   "14_DQ_Data_24PF2" : Bool = PLC "14_DQ_Data".24PF2 AT %DB1.DBX0.0, 1 s
   "19_AUTO_CMNDS_Data_PIT402_Target" : Real = PLC "19_AUTO_CMNDS_Data".PIT402_Target AT %DB1.DBD0, 1 s
   "80_From_HMI_RST_E500A_RT" : Bool = PLC "80_From_HMI".RST_E500A_RT AT %DB1.DBX0.0, 1 s
   "10_DI_Data_CV312_OPN" : Bool = PLC "10_DI_Data".CV312_OPN AT %DB1.DBX0.0, 1 s
   "10_DI_Data_CV312_CLSD" : Bool = PLC "10_DI_Data".CV312_CLSD AT %DB1.DBX0.0, 1 s
   "Clock_1Hz" : Bool = PLC Clock_1Hz AT %M0.5, 500 ms
   "14_DQ_Data_24K3(1)" : Bool = PLC "14_DQ_Data".24K3 AT %DB1.DBX0.0, 1 s
   "12_AI_Data_LIT305_SCALED" : Real = PLC "12_AI_Data".LIT305_SCALED AT %DB1.DBX0.0, 1 s
   "80_From_HMI_BWT_BYPASS(1)" : Bool = PLC "80_From_HMI".BWT_BYPASS AT %DB1.DBX0.0, 1 s
   "80_From_HMI_CRG_BLNK_MODE(1)" : Bool = PLC "80_From_HMI".CRG_BLNK_MODE AT %DB1.DBX0.0, 1 s
   "80_From_HMI_BWT_BYPASS" : Bool = PLC "80_From_HMI".BWT_BYPASS AT %DB1.DBX0.0, 1 s
   "80_From_HMI_CRG_BLNK_MODE" : Bool = PLC "80_From_HMI".CRG_BLNK_MODE AT %DB1.DBX0.0, 1 s
   "10_DI_Data_CV431_OPN" : Bool = PLC "10_DI_Data".CV431_OPN AT %DB1.DBX0.0, 1 s
   "10_DI_Data_CV431_CLSD" : Bool = PLC "10_DI_Data".CV431_CLSD AT %DB1.DBX0.0, 1 s
   "10_DI_Data_CV432_OPN" : Bool = PLC "10_DI_Data".CV432_OPN AT %DB1.DBX0.0, 1 s
   "10_DI_Data_CV432_CLSD" : Bool = PLC "10_DI_Data".CV432_CLSD AT %DB1.DBX0.0, 1 s
   "12_AI_Data_AT_O2_01_SCALED" : Real = PLC "12_AI_Data".AT_O2_01_SCALED AT %DB1.DBX0.0, 1 s
   "12_AI_Data_AT_O2_02_SCALED" : Real = PLC "12_AI_Data".AT_O2_02_SCALED AT %DB1.DBX0.0, 1 s
   "84_Setpoints_PIT102_Pilot_LowLow" : Real = PLC "84_Setpoints".PIT102_Pilot_LowLow AT %DB1.DBX0.0, 1 s
   "84_Setpoints_PIT102_Pilot_Low" : Real = PLC "84_Setpoints".PIT102_Pilot_Low AT %DB1.DBX0.0, 1 s
   "84_Setpoints_PIT102_Pilot_High" : Real = PLC "84_Setpoints".PIT102_Pilot_High AT %DB1.DBD0, 1 s
   "84_Setpoints_PIT102_Pilot_HighHigh" : Real = PLC "84_Setpoints".PIT102_Pilot_HighHigh AT %DB1.DBD0, 1 s
   "84_Setpoints_PIT102_Main_LowLow" : Real = PLC "84_Setpoints".PIT102_Main_LowLow AT %DB1.DBD0, 1 s
   "84_Setpoints_PIT102_Main_Low" : Real = PLC "84_Setpoints".PIT102_Main_Low AT %DB1.DBD0, 1 s
   "84_Setpoints_PIT102_Main_High" : Real = PLC "84_Setpoints".PIT102_Main_High AT %DB1.DBD0, 1 s
   "84_Setpoints_PIT102_Main_HighHigh" : Real = PLC "84_Setpoints".PIT102_Main_HighHigh AT %DB1.DBD0, 1 s
   "84_Setpoints_TIT401_High" : Real = PLC "84_Setpoints".TIT401_High AT %DB1.DBD0, 1 s
   "84_Setpoints_TIT401_HighHigh" : Real = PLC "84_Setpoints".TIT401_HighHigh AT %DB1.DBD0, 1 s
   "84_Setpoints_PIT402_Pilot_LowLow" : Real = PLC "84_Setpoints".PIT402_Pilot_LowLow AT %DB1.DBD0, 1 s
   "84_Setpoints_PIT402_Pilot_Low" : Real = PLC "84_Setpoints".PIT402_Pilot_Low AT %DB1.DBD0, 1 s
   "84_Setpoints_PIT402_Pilot_High" : Real = PLC "84_Setpoints".PIT402_Pilot_High AT %DB1.DBD0, 1 s
   "84_Setpoints_PIT402_Pilot_HighHigh" : Real = PLC "142_P304_HRS_RUN_DB".HRS AT %DB1.DBD0, 1 s
   "84_Setpoints_PIT402_Main_LowLow" : Real = PLC "84_Setpoints".PIT402_Main_LowLow AT %DB1.DBD0, 1 s
   "84_Setpoints_PIT402_Main_Low" : Real = PLC "84_Setpoints".PIT402_Main_Low AT %DB1.DBD0, 1 s
   "84_Setpoints_PIT402_Main_High" : Real = PLC "84_Setpoints".PIT402_Main_High AT %DB1.DBD0, 1 s
   "84_Setpoints_PIT402_Main_HighHigh" : Real = PLC "84_Setpoints".PIT402_Main_HighHigh AT %DB1.DBD0, 1 s
   "84_Setpoints_PIT112_LowLow" : Real = PLC "84_Setpoints".PIT112_LowLow AT %DB1.DBD0, 1 s
   "84_Setpoints_PIT112_Low" : Real = PLC "84_Setpoints".PIT112_Low AT %DB1.DBD0, 1 s
   "84_Setpoints_PIT112_High" : Real = PLC "84_Setpoints".PIT112_High AT %DB1.DBD0, 1 s
   "84_Setpoints_PIT112_HighHigh" : Real = PLC "84_Setpoints".PIT112_HighHigh AT %DB1.DBD0, 1 s
   "84_Setpoints_TIT315_High" : Real = PLC "84_Setpoints".TIT315_High AT %DB1.DBX0.0, 1 s
   "84_Setpoints_TIT315_HighHigh" : Real = PLC "84_Setpoints".TIT315_HighHigh AT %DB1.DBD0, 1 s
   "84_Setpoints_TIT319_High" : Real = PLC "84_Setpoints".TIT319_High AT %DB1.DBD0, 1 s
   "84_Setpoints_TIT319_HighHigh" : Real = PLC "84_Setpoints".TIT319_HighHigh AT %DB1.DBD0, 1 s
   "84_Setpoints_TIT360_High" : Real = PLC "84_Setpoints".TIT360_High AT %DB1.DBD0, 1 s
   "84_Setpoints_TIT360_HighHigh" : Real = PLC "84_Setpoints".TIT360_HighHigh AT %DB1.DBD0, 1 s
   "84_Setpoints_PIT359_LowLow" : Real = PLC "84_Setpoints".PIT359_LowLow AT %DB1.DBD0, 1 s
   "84_Setpoints_PIT359_Low" : Real = PLC "84_Setpoints".PIT359_Low AT %DB1.DBD0, 1 s
   "84_Setpoints_PIT359_High" : Real = PLC "84_Setpoints".PIT359_High AT %DB1.DBD0, 1 s
   "84_Setpoints_PIT359_HighHigh" : Real = PLC "84_Setpoints".PIT359_HighHigh AT %DB1.DBD0, 1 s
   "84_Setpoints_PIT316_LowLow" : Real = PLC "84_Setpoints".PIT316_LowLow AT %DB1.DBD0, 1 s
   "84_Setpoints_PIT316_Low" : Real = PLC "84_Setpoints".PIT316_Low AT %DB1.DBD0, 1 s
   "84_Setpoints_PIT316_High" : Real = PLC "84_Setpoints".PIT316_High AT %DB1.DBD0, 1 s
   "84_Setpoints_PIT316_HighHigh" : Real = PLC "84_Setpoints".PIT316_HighHigh AT %DB1.DBD0, 1 s
   "14_DQ_Data_CV431_432_CNTRL" : Bool = PLC "14_DQ_Data".CV431_432_CNTRL AT %DB1.DBX0.0, 1 s
   "14_DQ_Data_R2_SPR_DQ_0_7" : Bool = PLC "14_DQ_Data".R2_SPR_DQ_0_7 AT %DB1.DBX0.0, 1 s
   "14_DQ_Data_R2_SPR_DQ_1_0" : Bool = PLC "14_DQ_Data".R2_SPR_DQ_1_0 AT %DB1.DBX0.0, 1 s
   "80_From_HMI_MAN_DQ_0_0" : Bool = PLC "80_From_HMI".MAN_DQ_0_0 AT %DB1.DBX0.0, 1 s
   "80_From_HMI_MAN_DQ_0_1" : Bool = PLC "80_From_HMI".MAN_DQ_0_1 AT %DB1.DBX0.0, 1 s
   "80_From_HMI_MAN_DQ_0_2" : Bool = PLC "80_From_HMI".MAN_DQ_0_2 AT %DB1.DBX0.0, 1 s
   "80_From_HMI_MAN_DQ_0_3" : Bool = PLC "80_From_HMI".MAN_DQ_0_3 AT %DB1.DBX0.0, 1 s
   "80_From_HMI_MAN_DQ_0_4" : Bool = PLC "80_From_HMI".MAN_DQ_0_4 AT %DB1.DBX0.0, 1 s
   "80_From_HMI_MAN_DQ_0_5" : Bool = PLC "80_From_HMI".MAN_DQ_0_5 AT %DB1.DBX0.0, 1 s
   "80_From_HMI_MAN_DQ_0_6" : Bool = PLC "80_From_HMI".MAN_DQ_0_6 AT %DB1.DBX0.0, 1 s
   "80_From_HMI_MAN_DQ_0_7(1)" : Bool = PLC "80_From_HMI".MAN_DQ_0_7 AT %DB1.DBX0.0, 1 s
   "80_From_HMI_MAN_DQ_1_0(1)" : Bool = PLC "80_From_HMI".MAN_DQ_1_0 AT %DB1.DBX0.0, 1 s
   "80_From_HMI_MAN_DQ_1_1" : Bool = PLC "80_From_HMI".MAN_DQ_1_1 AT %DB1.DBX0.0, 1 s
   "80_From_HMI_MAN_DQ_1_2" : Bool = PLC "80_From_HMI".MAN_DQ_1_2 AT %DB1.DBX0.0, 1 s
   "80_From_HMI_MAN_DQ_1_3" : Bool = PLC "80_From_HMI".MAN_DQ_1_3 AT %DB1.DBX0.0, 1 s
   "80_From_HMI_MAN_DQ_1_4" : Bool = PLC "80_From_HMI".MAN_DQ_1_4 AT %DB1.DBX0.0, 1 s
   "80_From_HMI_MAN_DQ_1_5" : Bool = PLC "80_From_HMI".MAN_DQ_1_5 AT %DB1.DBX0.0, 1 s
   "80_From_HMI_MAN_DQ_1_6(1)" : Bool = PLC "80_From_HMI".MAN_DQ_1_6 AT %DB1.DBX0.0, 1 s
   "80_From_HMI_MAN_DQ_1_7" : Bool = PLC "80_From_HMI".MAN_DQ_1_7 AT %DB1.DBX0.0, 1 s
   "10_DI_Data_E139_READY" : Bool = PLC "10_DI_Data".E139_READY AT %DB1.DBX0.0, 1 s
   "10_DI_Data_E139_RUNNING(1)" : Bool = PLC "10_DI_Data".E139_RUNNING AT %DB1.DBX0.0, 1 s
   "10_DI_Data_E139_VSD_FLT" : Bool = PLC "10_DI_Data".E139_VSD_FLT AT %DB1.DBX0.0, 1 s
   "10_DI_Data_MCCP_5PG1_OK" : Bool = PLC "10_DI_Data".MCCP_5PG1_OK AT %DB1.DBX0.0, 1 s
   "10_DI_Data_R1_SPR_DI_3_7" : Bool = PLC "10_DI_Data".R1_SPR_DI_3_7 AT %DB1.DBX0.0, 1 s
   "84_Setpoints_AT_O2_1_Low" : Real = PLC "84_Setpoints".AT_O2_1_Low AT %DB1.DBD0, 1 s
   "84_Setpoints_PIT402_Main_Target" : Real = PLC "84_Setpoints".PIT402_Main_Target AT %DB1.DBX0.0, 1 s
   "84_Setpoints_PIT402_Pilot_Target" : Real = PLC "84_Setpoints".PIT402_Pilot_Target AT %DB1.DBD0, 1 s
   "14_DQ_Data_E139_CNTRL" : Bool = PLC RIO6_SPR_DI_63_7 AT %DB1.DBX0.0, 1 s
   "80_From_HMI_E139_SET_SPEED" : Real = PLC "80_From_HMI".E139_SET_SPEED AT %DB1.DBX0.0, 1 s
   "10_DI_Data_CV311_OPN(1)" : Bool = PLC "10_DI_Data".CV311_OPN AT %DB1.DBX0.0, 1 s
   "80_From_HMI_MAX_E500_RT" : LTime = PLC "80_From_HMI".MAX_E500_RT AT %DB1.DBX0.0, 1 s
   "68_Sys_Status_Data_IA_PRES_IN_RNG(1)" : Bool = PLC "68_Sys_Status_Data".IA_PRES_IN_RNG AT %DB1.DBX0.0, 1 s
   "68_Sys_Status_Data_FUEL_PRES_IN_RNG(1)" : Bool = PLC "68_Sys_Status_Data".FUEL_PRES_IN_RNG AT %DB1.DBX0.0, 1 s
   "16_AQ_Data_E139_SPEED" : Real = PLC "16_AQ_Data".E139_SPEED AT %DB1.DBD0, 1 s
   "16_AQ_Data_R1_SPR_AQ_102" : Real = PLC "16_AQ_Data".R1_SPR_AQ_102 AT %DB1.DBD0, 1 s
   "16_AQ_Data_R1_SPR_AQ_104" : Real = PLC "16_AQ_Data".R1_SPR_AQ_104 AT %DB1.DBD0, 1 s
   "80_From_HMI_MAN_AQ_INC_98(1)" : Bool = PLC "80_From_HMI".MAN_AQ_INC_98 AT %DB1.DBX0.0, 1 s
   "80_From_HMI_MAN_AQ_DEC_98(1)" : Bool = PLC "80_From_HMI".MAN_AQ_DEC_98 AT %DB1.DBX0.0, 1 s
   "80_From_HMI_MAN_AQ_INC_100" : Bool = PLC "80_From_HMI".MAN_AQ_INC_100 AT %DB1.DBX0.0, 1 s
   "80_From_HMI_MAN_AQ_DEC_100" : Bool = PLC "80_From_HMI".MAN_AQ_DEC_100 AT %DB1.DBX0.0, 1 s
   "80_From_HMI_MAN_AQ_INC_102(1)" : Bool = PLC "80_From_HMI".MAN_AQ_INC_102 AT %DB1.DBX0.0, 1 s
   "80_From_HMI_MAN_AQ_DEC_102(1)" : Bool = PLC "80_From_HMI".MAN_AQ_DEC_102 AT %DB1.DBX0.0, 1 s
   "80_From_HMI_MAN_AQ_DEC_104" : Bool = PLC "80_From_HMI".MAN_AQ_DEC_104 AT %DB1.DBX0.0, 1 s
   "80_From_HMI_MAN_AQ_INC_104" : Bool = PLC "80_From_HMI".MAN_AQ_INC_104 AT %DB1.DBX0.0, 1 s
   "80_From_HMI_STOP_IGG" : Bool = PLC "80_From_HMI".STOP_IGG AT %DB1.DBX0.0, 1 s
   "80_From_HMI_Request_Auto(1)" : Bool = PLC "80_From_HMI".Request_Auto AT %DB1.DBX0.0, 1 s
   "80_From_HMI_RST_AUT_SEQ(1)" : Bool = PLC "80_From_HMI".RST_AUT_SEQ AT %DB1.DBX0.0, 1 s
   "80_From_HMI_FAT_Mode" : Bool = PLC "80_From_HMI".FAT_Mode AT %DB1.DBX0.0, 1 s
   "80_From_HMI_IGG_STND_ALN" : Bool = PLC "80_From_HMI".IGG_STND_ALN AT %DB1.DBX0.0, 1 s
   "80_From_HMI_P301_PRSNT(1)" : Bool = PLC "80_From_HMI".P301_PRSNT AT %DB1.DBX0.0, 1 s
   "80_From_HMI_CV312_PRSNT" : Bool = PLC "80_From_HMI".CV312_PRSNT AT %DB1.DBX0.0, 1 s
   "80_From_HMI_CV431_PRSNT" : Bool = PLC "80_From_HMI".CV431_PRSNT AT %DB1.DBX0.0, 1 s
   "80_From_HMI_CV432_PRSNT" : Bool = PLC "80_From_HMI".CV432_PRSNT AT %DB1.DBX0.0, 1 s
   "80_From_HMI_SLNCE_BZR" : Bool = PLC "80_From_HMI".SLNCE_BZR AT %DB1.DBX0.0, 1 s
   "84_Setpoints_PIT102_Post_LowLow" : Real = PLC "84_Setpoints".PIT102_Post_LowLow AT %DB1.DBD0, 1 s
   "84_Setpoints_PIT102_Post_Low" : Real = PLC "84_Setpoints".PIT102_Post_Low AT %DB1.DBD0, 1 s
   "84_Setpoints_PIT102_Post_HighHigh" : Real = PLC "84_Setpoints".PIT102_Post_HighHigh AT %DB1.DBD0, 1 s
   "84_Setpoints_PIT102_Post_High" : Real = PLC "84_Setpoints".PIT102_Post_High AT %DB1.DBD0, 1 s
   "12_AI_Data_R1_SPR_AI_126_SCALED" : Real = PLC "12_AI_Data".R1_SPR_AI_126_SCALED AT %DB1.DBX0.0, 1 s
   "12_AI_Data_R1_SPR_AI_132_SCALED" : Real = PLC "12_AI_Data".R1_SPR_AI_132_SCALED AT %DB1.DBD0, 1 s
   "84_Setpoints_PIT402_Post_High" : Real = PLC "84_Setpoints".PIT402_Post_High AT %DB1.DBD0, 1 s
   "84_Setpoints_PIT402_Post_HighHigh" : Real = PLC "84_Setpoints".PIT402_Post_HighHigh AT %DB1.DBD0, 1 s
   "84_Setpoints_PIT402_Post_Low" : Real = PLC "84_Setpoints".PIT402_Post_Low AT %DB1.DBD0, 1 s
   "84_Setpoints_PIT402_Post_LowLow" : Real = PLC "84_Setpoints".PIT402_Post_LowLow AT %DB1.DBD0, 1 s
   "84_Setpoints_PIT402_Pilot_Target(1)" : Real = PLC "84_Setpoints".PIT402_Pilot_Target AT %DB1.DBD0, 1 s
   "84_Setpoints_PIT402_Main_Target(1)" : Real = PLC "84_Setpoints".PIT402_Main_Target AT %DB1.DBD0, 1 s
   "84_Setpoints_PIT402_Post_Target_Start" : Real = PLC "84_Setpoints".PIT402_Post_Target_Start AT %DB1.DBD0, 1 s
   "84_Setpoints_PIT401_Post_Target_Max" : Real = PLC "84_Setpoints".PIT401_Post_Target_Max AT %DB1.DBD0, 1 s
   "86_Times_PRE_BC_STRT_CMND_DLY" : Time = PLC "86_Times".PRE_BC_STRT_CMND_DLY AT %DB1.DBD0, 1 s
   "86_Times_PRE_CV203_CLS_CMND_DLY" : Time = PLC "86_Times".PRE_CV203_CLS_CMND_DLY AT %DB1.DBD0, 1 s
   "86_Times_POST_P301_STOP_DLY" : Time = PLC "86_Times".POST_P301_STOP_DLY AT %DB1.DBD0, 1 s
   "86_Times_POST_CV311_CLS_DLY" : Time = PLC "86_Times".POST_CV311_CLS_DLY AT %DB1.DBD0, 1 s
   "86_Times_POST_CV321_OPN_DLY" : Time = PLC "86_Times".POST_CV321_OPN_DLY AT %DB1.DBD0, 1 s
   "86_Times_CV311_MAX_TRVL_TIME" : Time = PLC "86_Times".CV311_MAX_TRVL_TIME AT %DB1.DBD0, 1 s
   "86_Times_CV312_MAX_TRVL_TIME" : Time = PLC "86_Times".CV312_MAX_TRVL_TIME AT %DB1.DBD0, 1 s
   "86_Times_CV321_MAX_TRVL_TIME" : Time = PLC "86_Times".CV321_MAX_TRVL_TIME AT %DB1.DBD0, 1 s
   "86_Times_CV322_MAX_TRVL_TIME" : Time = PLC "86_Times".CV322_MAX_TRVL_TIME AT %DB1.DBD0, 1 s
   "86_Times_CV401_MAX_TRVL_TIME" : Time = PLC "86_Times".CV401_MAX_TRVL_TIME AT %DB1.DBD0, 1 s
   "86_Times_CV431_MAX_TRVL_TIME" : Time = PLC "86_Times".CV431_MAX_TRVL_TIME AT %DB1.DBD0, 1 s
   "86_Times_CV432_MAX_TRVL_TIME" : Time = PLC "86_Times".CV432_MAX_TRVL_TIME AT %DB1.DBD0, 1 s
   "86_Times_STEP_MAX_TIME_STP_001(2)" : Time = PLC "86_Times".STEP_MAX_TIME_STP_001 AT %DB1.DBW0, 1 s
   "86_Times_STEP_MAX_TIME_STP_005(2)" : Time = PLC "86_Times".STEP_MAX_TIME_STP_005 AT %DB1.DBW0, 1 s
   "86_Times_STEP_MAX_TIME_STP_010(2)" : Time = PLC "86_Times".STEP_MAX_TIME_STP_010 AT %DB1.DBW0, 1 s
   "86_Times_STEP_MAX_TIME_STP_020(2)" : Time = PLC "86_Times".STEP_MAX_TIME_STP_020 AT %DB1.DBW0, 1 s
   "86_Times_STEP_MAX_TIME_STP_030(2)" : Time = PLC "86_Times".STEP_MAX_TIME_STP_030 AT %DB1.DBW0, 1 s
   "86_Times_STEP_MAX_TIME_STP_040(2)" : Time = PLC "86_Times".STEP_MAX_TIME_STP_040 AT %DB1.DBW0, 1 s
   "86_Times_STEP_MAX_TIME_STP_050(2)" : Time = PLC "86_Times".STEP_MAX_TIME_STP_050 AT %DB1.DBW0, 1 s
   "86_Times_STEP_MAX_TIME_STP_060(2)" : Time = PLC "86_Times".STEP_MAX_TIME_STP_060 AT %DB1.DBW0, 1 s
   "86_Times_STEP_MAX_TIME_STP_070(2)" : Time = PLC "86_Times".STEP_MAX_TIME_STP_070 AT %DB1.DBW0, 1 s
   "86_Times_STEP_MAX_TIME_STP_080(2)" : Time = PLC "86_Times".STEP_MAX_TIME_STP_080 AT %DB1.DBW0, 1 s
   "86_Times_STEP_MAX_TIME_STP_090(2)" : Time = PLC "86_Times".STEP_MAX_TIME_STP_090 AT %DB1.DBW0, 1 s
   "86_Times_STEP_MAX_TIME_STP_100(2)" : Time = PLC "86_Times".STEP_MAX_TIME_STP_100 AT %DB1.DBW0, 1 s
   "86_Times_STEP_MAX_TIME_STP_110(2)" : Time = PLC "86_Times".STEP_MAX_TIME_STP_110 AT %DB1.DBW0, 1 s
   "86_Times_STEP_MAX_TIME_STP_120(2)" : Time = PLC "86_Times".STEP_MAX_TIME_STP_120 AT %DB1.DBW0, 1 s
   "86_Times_STEP_MAX_TIME_STP_130(2)" : Time = PLC "86_Times".STEP_MAX_TIME_STP_130 AT %DB1.DBW0, 1 s
   "86_Times_STEP_MAX_TIME_STP_140(2)" : Time = PLC "86_Times".STEP_MAX_TIME_STP_140 AT %DB1.DBW0, 1 s
   "86_Times_STEP_MAX_TIME_STP_150(2)" : Time = PLC "86_Times".STEP_MAX_TIME_STP_150 AT %DB1.DBW0, 1 s
   "86_Times_STEP_MAX_TIME_STP_160(2)" : Time = PLC "86_Times".STEP_MAX_TIME_STP_160 AT %DB1.DBW0, 1 s
   "86_Times_STEP_MAX_TIME_STP_170(2)" : Time = PLC "86_Times".STEP_MAX_TIME_STP_170 AT %DB1.DBW0, 1 s
   "86_Times_STEP_MAX_TIME_STP_180(2)" : Time = PLC "86_Times".STEP_MAX_TIME_STP_180 AT %DB1.DBW0, 1 s
   "86_Times_STEP_MAX_TIME_STP_190(2)" : Time = PLC "86_Times".STEP_MAX_TIME_STP_190 AT %DB1.DBW0, 1 s
   "86_Times_STEP_MAX_TIME_STP_200(2)" : Time = PLC "86_Times".STEP_MAX_TIME_STP_200 AT %DB1.DBW0, 1 s
   "86_Times_STEP_MAX_TIME_STP_210(2)" : Time = PLC "86_Times".STEP_MAX_TIME_STP_210 AT %DB1.DBW0, 1 s
   "86_Times_STEP_MAX_TIME_STP_220(2)" : Time = PLC "86_Times".STEP_MAX_TIME_STP_220 AT %DB1.DBW0, 1 s
   "86_Times_STEP_MAX_TIME_STP_230(2)" : Time = PLC "86_Times".STEP_MAX_TIME_STP_230 AT %DB1.DBW0, 1 s
   "86_Times_STEP_MAX_TIME_STP_240(2)" : Time = PLC "86_Times".STEP_MAX_TIME_STP_240 AT %DB1.DBW0, 1 s
   "86_Times_STEP_MAX_TIME_STP_250(2)" : Time = PLC "86_Times".STEP_MAX_TIME_STP_250 AT %DB1.DBW0, 1 s
   "86_Times_STEP_MAX_TIME_STP_260(2)" : Time = PLC "86_Times".STEP_MAX_TIME_STP_260 AT %DB1.DBW0, 1 s
   "86_Times_STEP_MAX_TIME_STP_270(2)" : Time = PLC "86_Times".STEP_MAX_TIME_STP_270 AT %DB1.DBW0, 1 s
   "86_Times_STEP_MAX_TIME_STP_280(2)" : Time = PLC "86_Times".STEP_MAX_TIME_STP_280 AT %DB1.DBW0, 1 s
   "86_Times_STEP_MAX_TIME_STP_290(2)" : Time = PLC "86_Times".STEP_MAX_TIME_STP_290 AT %DB1.DBW0, 1 s
   "86_Times_STEP_MAX_TIME_STP_300(2)" : Time = PLC "86_Times".STEP_MAX_TIME_STP_300 AT %DB1.DBW0, 1 s
   "86_Times_STEP_MAX_TIME_STP_310(2)" : Time = PLC "86_Times".STEP_MAX_TIME_STP_310 AT %DB1.DBW0, 1 s
   "86_Times_STEP_MAX_TIME_STP_320(2)" : Time = PLC "86_Times".STEP_MAX_TIME_STP_320 AT %DB1.DBW0, 1 s
   "86_Times_STEP_MAX_TIME_STP_330(2)" : Time = PLC "86_Times".STEP_MAX_TIME_STP_330 AT %DB1.DBW0, 1 s
   "86_Times_STEP_MAX_TIME_STP_340(2)" : Time = PLC "86_Times".STEP_MAX_TIME_STP_340 AT %DB1.DBW0, 1 s
   "86_Times_STEP_MAX_TIME_STP_350(2)" : Time = PLC "86_Times".STEP_MAX_TIME_STP_350 AT %DB1.DBW0, 1 s
   "86_Times_STEP_MAX_TIME_STP_360(2)" : Time = PLC "86_Times".STEP_MAX_TIME_STP_360 AT %DB1.DBW0, 1 s
   "86_Times_STEP_MAX_TIME_STP_370(2)" : Time = PLC "86_Times".STEP_MAX_TIME_STP_370 AT %DB1.DBW0, 1 s
   "86_Times_STEP_MAX_TIME_STP_380(2)" : Time = PLC "86_Times".STEP_MAX_TIME_STP_380 AT %DB1.DBW0, 1 s
   "86_Times_STEP_MAX_TIME_STP_390(2)" : Time = PLC "86_Times".STEP_MAX_TIME_STP_390 AT %DB1.DBW0, 1 s
   "86_Times_STEP_MAX_TIME_STP_400(2)" : Time = PLC "86_Times".STEP_MAX_TIME_STP_400 AT %DB1.DBW0, 1 s
   "86_Times_STEP_MAX_TIME_STP_410(2)" : Time = PLC "86_Times".STEP_MAX_TIME_STP_410 AT %DB1.DBW0, 1 s
   "86_Times_STEP_MAX_TIME_STP_420(2)" : Time = PLC TT426_FPT_ALM_ANALOG_DB."LOW LEVEL VALUE (L)" AT %DB1.DBW0, 1 s
   "86_Times_STEP_MAX_TIME_STP_430(2)" : Time = PLC "86_Times".STEP_MAX_TIME_STP_430 AT %DB1.DBW0, 1 s
   "86_Times_STEP_MAX_TIME_STP_440(2)" : Time = PLC "86_Times".STEP_MAX_TIME_STP_440 AT %DB1.DBW0, 1 s
   "86_Times_STEP_MAX_TIME_STP_450(2)" : Time = PLC "86_Times".STEP_MAX_TIME_STP_450 AT %DB1.DBW0, 1 s
   "86_Times_STEP_MAX_TIME_STP_460(2)" : Time = PLC "86_Times".STEP_MAX_TIME_STP_460 AT %DB1.DBW0, 1 s
   "86_Times_STEP_MAX_TIME_STP_470(2)" : Time = PLC "86_Times".STEP_MAX_TIME_STP_470 AT %DB1.DBW0, 1 s
   "86_Times_STEP_MAX_TIME_STP_480(2)" : Time = PLC "86_Times".STEP_MAX_TIME_STP_480 AT %DB1.DBW0, 1 s
   "86_Times_STEP_MAX_TIME_STP_490(2)" : Time = PLC "86_Times".STEP_MAX_TIME_STP_490 AT %DB1.DBW0, 1 s
   "86_Times_STEP_MAX_TIME_STP_500(2)" : Time = PLC "86_Times".STEP_MAX_TIME_STP_500 AT %DB1.DBW0, 1 s
   "Logging SD Card Overflow" : Bool AT %DB1.DBX0.0
      on ChangeValue: "SD_Card_Overflow"()
   "CSW_Animation_DB_Animation" : Int = PLC CSW_Animation_DB.Animation, 1 s
   "504_Tank Grouping_DB2020_Time Left Tank_Time Left m Tank 1" : DInt = PLC "504_Tank Grouping_DB2020"."Time Left Tank"."Time Left m Tank 1", 1 s
   "504_Tank Grouping_DB2020_Time Left Tank_Time Left h Tank 1" : DInt = PLC "504_Tank Grouping_DB2020"."Time Left Tank"."Time Left h Tank 1", 1 s
   "504_Tank Grouping_DB2020_Time Left Tank_Time Left d Tank 1" : DInt = PLC "504_Tank Grouping_DB2020"."Time Left Tank"."Time Left d Tank 1", 1 s
   "504_Tank Grouping_DB2020_Time Left Tank_Time Left m Tank 2" : DInt = PLC "504_Tank Grouping_DB2020"."Time Left Tank"."Time Left m Tank 2", 1 s
   "504_Tank Grouping_DB2020_Time Left Tank_Time Left h Tank 14" : DInt = PLC "504_Tank Grouping_DB2020"."Time Left Tank"."Time Left h Tank 14", 1 s
   "504_Tank Grouping_DB2020_Time Left Tank_Time Left d Tank 14" : DInt = PLC "504_Tank Grouping_DB2020"."Time Left Tank"."Time Left d Tank 14", 1 s
   "504_Tank Grouping_DB2020_Time Left Tank_Time Left m Tank 14" : DInt = PLC "504_Tank Grouping_DB2020"."Time Left Tank"."Time Left m Tank 14", 1 s
   "504_Tank Grouping_DB2020_Time Left Tank_Time Left h Tank 2" : DInt = PLC "504_Tank Grouping_DB2020"."Time Left Tank"."Time Left h Tank 2", 1 s
   "504_Tank Grouping_DB2020_Time Left Tank_Time Left d Tank 2" : DInt = PLC "504_Tank Grouping_DB2020"."Time Left Tank"."Time Left d Tank 2", 1 s
   "504_Tank Grouping_DB2020_Time Left Tank_Time Left m Tank 3" : DInt = PLC "504_Tank Grouping_DB2020"."Time Left Tank"."Time Left m Tank 3", 1 s
   "504_Tank Grouping_DB2020_Time Left Tank_Time Left h Tank 3" : DInt = PLC "504_Tank Grouping_DB2020"."Time Left Tank"."Time Left h Tank 3", 1 s
   "504_Tank Grouping_DB2020_Time Left Tank_Time Left d Tank 3" : DInt = PLC "504_Tank Grouping_DB2020"."Time Left Tank"."Time Left d Tank 3", 1 s
   "504_Tank Grouping_DB2020_Time Left Tank_Time Left m Tank 4" : DInt = PLC "504_Tank Grouping_DB2020"."Time Left Tank"."Time Left m Tank 4", 1 s
   "504_Tank Grouping_DB2020_Time Left Tank_Time Left h Tank 4" : DInt = PLC "504_Tank Grouping_DB2020"."Time Left Tank"."Time Left h Tank 4", 1 s
   "504_Tank Grouping_DB2020_Time Left Tank_Time Left d Tank 4" : DInt = PLC "504_Tank Grouping_DB2020"."Time Left Tank"."Time Left d Tank 4", 1 s
   "504_Tank Grouping_DB2020_Time Left Tank_Time Left m Tank 5" : DInt = PLC "504_Tank Grouping_DB2020"."Time Left Tank"."Time Left m Tank 5", 1 s
   "504_Tank Grouping_DB2020_Time Left Tank_Time Left h Tank 5" : DInt = PLC "504_Tank Grouping_DB2020"."Time Left Tank"."Time Left h Tank 5", 1 s
   "504_Tank Grouping_DB2020_Time Left Tank_Time Left d Tank 5" : DInt = PLC "504_Tank Grouping_DB2020"."Time Left Tank"."Time Left d Tank 5", 1 s
   "504_Tank Grouping_DB2020_Time Left Tank_Time Left m Tank 6" : DInt = PLC "504_Tank Grouping_DB2020"."Time Left Tank"."Time Left m Tank 6", 1 s
   "504_Tank Grouping_DB2020_Time Left Tank_Time Left h Tank 6" : DInt = PLC "504_Tank Grouping_DB2020"."Time Left Tank"."Time Left h Tank 6", 1 s
   "504_Tank Grouping_DB2020_Time Left Tank_Time Left d Tank 6" : DInt = PLC "504_Tank Grouping_DB2020"."Time Left Tank"."Time Left d Tank 6", 1 s
   "504_Tank Grouping_DB2020_Time Left Tank_Time Left m Tank 7" : DInt = PLC "504_Tank Grouping_DB2020"."Time Left Tank"."Time Left m Tank 7", 1 s
   "504_Tank Grouping_DB2020_Time Left Tank_Time Left h Tank 7" : DInt = PLC "504_Tank Grouping_DB2020"."Time Left Tank"."Time Left h Tank 7", 1 s
   "504_Tank Grouping_DB2020_Time Left Tank_Time Left d Tank 7" : DInt = PLC "504_Tank Grouping_DB2020"."Time Left Tank"."Time Left d Tank 7", 1 s
   "504_Tank Grouping_DB2020_Time Left Tank_Time Left m Tank 8" : DInt = PLC "504_Tank Grouping_DB2020"."Time Left Tank"."Time Left m Tank 8", 1 s
   "504_Tank Grouping_DB2020_Time Left Tank_Time Left h Tank 8" : DInt = PLC "504_Tank Grouping_DB2020"."Time Left Tank"."Time Left h Tank 8", 1 s
   "504_Tank Grouping_DB2020_Time Left Tank_Time Left d Tank 8" : DInt = PLC "504_Tank Grouping_DB2020"."Time Left Tank"."Time Left d Tank 8", 1 s
   "504_Tank Grouping_DB2020_Time Left Tank_Time Left m Tank 9" : DInt = PLC "2062_Warning_Data"."Alarm Tank P6", 1 s
   "504_Tank Grouping_DB2020_Time Left Tank_Time Left h Tank 9" : DInt = PLC "504_Tank Grouping_DB2020"."Time Left Tank"."Time Left h Tank 9", 1 s
   "504_Tank Grouping_DB2020_Time Left Tank_Time Left d Tank 9" : DInt = PLC "504_Tank Grouping_DB2020"."Time Left Tank"."Time Left d Tank 9", 1 s
   "504_Tank Grouping_DB2020_Time Left Tank_Time Left m Tank 10" : DInt = PLC "504_Tank Grouping_DB2020"."Time Left Tank"."Time Left m Tank 10", 1 s
   "504_Tank Grouping_DB2020_Time Left Tank_Time Left h Tank 10" : DInt = PLC "504_Tank Grouping_DB2020"."Time Left Tank"."Time Left h Tank 10", 1 s
   "504_Tank Grouping_DB2020_Time Left Tank_Time Left d Tank 10" : DInt = PLC "504_Tank Grouping_DB2020"."Time Left Tank"."Time Left d Tank 10", 1 s
   "504_Tank Grouping_DB2020_Time Left Tank_Time Left m Tank 11" : DInt = PLC "504_Tank Grouping_DB2020"."Time Left Tank"."Time Left m Tank 11", 1 s
   "504_Tank Grouping_DB2020_Time Left Tank_Time Left h Tank 11" : DInt = PLC "504_Tank Grouping_DB2020"."Time Left Tank"."Time Left h Tank 11", 1 s
   "504_Tank Grouping_DB2020_Time Left Tank_Time Left d Tank 11" : DInt = PLC "504_Tank Grouping_DB2020"."Time Left Tank"."Time Left d Tank 11", 1 s
   "504_Tank Grouping_DB2020_Time Left Tank_Time Left m Tank 12" : DInt = PLC "504_Tank Grouping_DB2020"."Time Left Tank"."Time Left m Tank 12", 1 s
   "504_Tank Grouping_DB2020_Time Left Tank_Time Left h Tank 12" : DInt = PLC "504_Tank Grouping_DB2020"."Time Left Tank"."Time Left h Tank 12", 1 s
   "504_Tank Grouping_DB2020_Time Left Tank_Time Left d Tank 12" : DInt = PLC "504_Tank Grouping_DB2020"."Time Left Tank"."Time Left d Tank 12", 1 s
   "504_Tank Grouping_DB2020_Time Left Tank_Time Left m Tank 13" : DInt = PLC "504_Tank Grouping_DB2020"."Time Left Tank"."Time Left m Tank 13", 1 s
   "504_Tank Grouping_DB2020_Time Left Tank_Time Left h Tank 13" : DInt = PLC "504_Tank Grouping_DB2020"."Time Left Tank"."Time Left h Tank 13", 1 s
   "504_Tank Grouping_DB2020_Time Left Tank_Time Left d Tank 13" : DInt = PLC "504_Tank Grouping_DB2020"."Time Left Tank"."Time Left d Tank 13", 1 s

HMI tags "Warnings"
   "62_Warning_Data_BC_WARNING_WORD_01" : Word = PLC "62_Warning_Data".BC_WARNING_WORD_01 AT %DB62.DBW0, 1 s
   "62_Warning_Data_BC_WARNING_WORD_02" : Word = PLC "62_Warning_Data".BC_WARNING_WORD_02 AT %DB62.DBW2, 1 s
   "62_Warning_Data_BC_WARNING_WORD_03" : Word = PLC "62_Warning_Data".BC_WARNING_WORD_03 AT %DB62.DBW4, 1 s
   "62_Warning_Data_BC_WARNING_WORD_04" : Word = PLC "62_Warning_Data".BC_WARNING_WORD_04 AT %DB62.DBW6, 1 s
   "62_Warning_Data_BC_WARNING_WORD_05" : Word = PLC "62_Warning_Data".BC_WARNING_WORD_05 AT %DB62.DBW8, 1 s
   "62_Warning_Data_BC_WARNING_WORD_06" : Word = PLC "62_Warning_Data".BC_WARNING_WORD_06 AT %DB62.DBW10, 1 s
   "62_Warning_Data_IGG_WARNING_WORD_01" : Word = PLC "62_Warning_Data".IGG_WARNING_WORD_01 AT %DB62.DBW0, 1 s
   "62_Warning_Data_IGG_WARNING_WORD_02" : Word = PLC "62_Warning_Data".IGG_WARNING_WORD_02 AT %DB62.DBW2, 1 s
   "62_Warning_Data_IGG_WARNING_WORD_03" : Word = PLC "62_Warning_Data".IGG_WARNING_WORD_03 AT %DB62.DBW4, 1 s
   "62_Warning_Data_IGG_WARNING_WORD_04" : Word = PLC "62_Warning_Data".IGG_WARNING_WORD_04 AT %DB62.DBW6, 1 s
   "62_Warning_Data_IGG_WARNING_WORD_05" : Word = PLC "62_Warning_Data".IGG_WARNING_WORD_05 AT %DB62.DBW8, 1 s
   "62_Warning_Data_IGG_WARNING_WORD_06" : Word = PLC "62_Warning_Data".IGG_WARNING_WORD_06 AT %DB62.DBW10, 1 s

